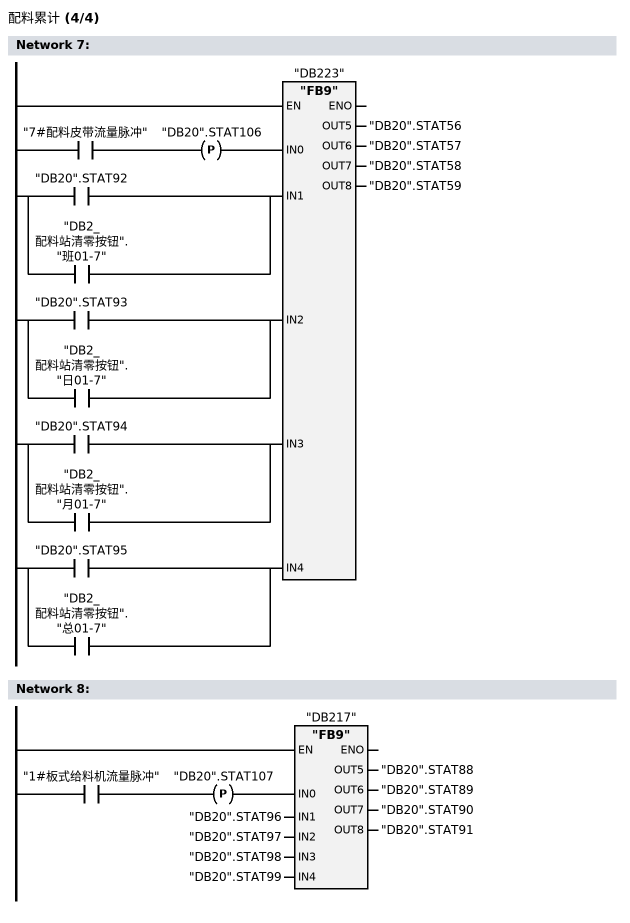
   RUNG wire#powerrail
      "DB223"(IN0 := wire#w1, IN1 := wire#w2, IN2 := wire#w3, IN3 := wire#w4, IN4 := wire#w5, OUT5 => "DB20".STAT56, OUT6 => "DB20".STAT57, OUT7 => "DB20".STAT58, OUT8 => "DB20".STAT59)
   END_RUNG
   RUNG wire#powerrail
      Contact( "7#配料皮带流量脉冲" )
      P_Trig( "DB20".STAT106 )
   END_RUNG wire#w1
   RUNG wire#powerrail
      Contact( "DB20".STAT92 )
   END_RUNG wire#w2
   RUNG wire#powerrail
      Contact( "DB2_配料站清零按钮"."班01-7" )
   END_RUNG wire#w2
   RUNG wire#powerrail
      Contact( "DB20".STAT93 )
   END_RUNG wire#w3
   RUNG wire#powerrail
      Contact( "DB2_配料站清零按钮"."日01-7" )
   END_RUNG wire#w3
   RUNG wire#powerrail
      Contact( "DB20".STAT94 )
   END_RUNG wire#w4
   RUNG wire#powerrail
      Contact( "DB2_配料站清零按钮"."月01-7" )
   END_RUNG wire#w4
   RUNG wire#powerrail
      Contact( "DB20".STAT95 )
   END_RUNG wire#w5
   RUNG wire#powerrail
      Contact( "DB2_配料站清零按钮"."总01-7" )
   END_RUNG wire#w5
   // the same network as SCL:
   #_w1 := "7#配料皮带流量脉冲" AND NOT "DB20".STAT106;   // rising edge
   "DB20".STAT106 := "7#配料皮带流量脉冲";
   "DB223"(IN0 := #_w1,   // "FB9"
           IN1 := "DB20".STAT92 OR "DB2_配料站清零按钮"."班01-7",
           IN2 := "DB20".STAT93 OR "DB2_配料站清零按钮"."日01-7",
           IN3 := "DB20".STAT94 OR "DB2_配料站清零按钮"."月01-7",
           IN4 := "DB20".STAT95 OR "DB2_配料站清零按钮"."总01-7",
           OUT5 => "DB20".STAT56,
           OUT6 => "DB20".STAT57,
           OUT7 => "DB20".STAT58,
           OUT8 => "DB20".STAT59);
END_REGION

REGION Network 8
   RUNG wire#powerrail
      "DB217"(IN0 := wire#w1, IN1 := "DB20".STAT96, IN2 := "DB20".STAT97, IN3 := "DB20".STAT98, IN4 := "DB20".STAT99, OUT5 => "DB20".STAT88, OUT6 => "DB20".STAT89, OUT7 => "DB20".STAT90, OUT8 => "DB20".STAT91)
   END_RUNG
   RUNG wire#powerrail
      Contact( "1#板式给料机流量脉冲" )
      P_Trig( "DB20".STAT107 )
   END_RUNG wire#w1
   // the same network as SCL:
   #_w1 := "1#板式给料机流量脉冲" AND NOT "DB20".STAT107;   // rising edge
   "DB20".STAT107 := "1#板式给料机流量脉冲";
   "DB217"(IN0 := #_w1,   // "FB9"
           IN1 := "DB20".STAT96,
           IN2 := "DB20".STAT97,
           IN3 := "DB20".STAT98,
           IN4 := "DB20".STAT99,
           OUT5 => "DB20".STAT88,
           OUT6 => "DB20".STAT89,
           OUT7 => "DB20".STAT90,
           OUT8 => "DB20".STAT91);
END_REGION
END_FUNCTION

FUNCTION "回转窑变频器驱动块" : Void   // FC111, LAD
{ S7_Optimized_Access := 'FALSE' }
VERSION : 0.1
   VAR_INPUT
      IN0 : Bool;   // IN0
      IN1 : Bool;   // IN1
      IN2 : Bool;   // IN2
      IN3 : Bool;   // IN3
      IN4 : Bool;   // IN4
      IN5 : Bool;   // IN5
      IN6 : Bool;   // IN6
      IN7 : Bool;   // IN7
      IN8 : Bool;   // IN8
   END_VAR
   VAR_IN_OUT
      OUT9 : Bool;   // OUT9
   END_VAR
BEGIN

REGION Network 1: OUT9
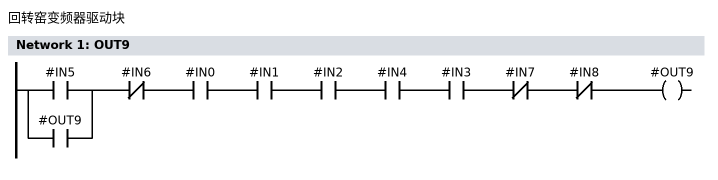
   RUNG wire#powerrail
      Contact( #IN5 )
      wire#w1
      I_Contact( #IN6 )
      Contact( #IN0 )
      Contact( #IN1 )
      Contact( #IN2 )
      Contact( #IN4 )
      Contact( #IN3 )
      I_Contact( #IN7 )
      I_Contact( #IN8 )
      Coil( #OUT9 )
   END_RUNG
   RUNG wire#powerrail
      Contact( #OUT9 )
   END_RUNG wire#w1
   // the same network as SCL:
   #OUT9 := (#IN5 OR #OUT9) AND NOT #IN6 AND #IN0 AND #IN1 AND #IN2 AND #IN4 AND #IN3 AND NOT #IN7 AND NOT #IN8;
END_REGION
END_FUNCTION

FUNCTION "回转窑接触器合闸块" : Void   // FC112, LAD
{ S7_Optimized_Access := 'FALSE' }
VERSION : 0.1
   VAR_INPUT
      IN0 : Bool;   // IN0
      IN1 : Bool;   // IN1
      IN2 : Bool;   // IN2
   END_VAR
   VAR_IN_OUT
      OUT3 : Bool;   // OUT3
   END_VAR
BEGIN

REGION Network 1: OUT3
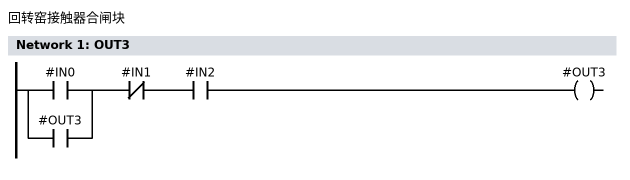
   RUNG wire#powerrail
      Contact( #IN0 )
      wire#w1
      I_Contact( #IN1 )
      Contact( #IN2 )
      Coil( #OUT3 )
   END_RUNG
   RUNG wire#powerrail
      Contact( #OUT3 )
   END_RUNG wire#w1
   // the same network as SCL:
   #OUT3 := (#IN0 OR #OUT3) AND NOT #IN1 AND #IN2;
END_REGION
END_FUNCTION

FUNCTION "稀油站功能块" : Void   // FC113, LAD
{ S7_Optimized_Access := 'FALSE' }
VERSION : 0.1
   VAR_INPUT
      LR1 : Bool;
      FAT1_1 : Bool;
      FAT1_2 : Bool;
      ST1 : Bool;
      STP1 : Bool;
      LR2 : Bool;
      FAT2_1 : Bool;
      FAT2_2 : Bool;
      ST2 : Bool;
      STP2 : Bool;
   END_VAR
   VAR_IN_OUT
      OUT10 : Bool;
      OUT11 : Bool;
   END_VAR
BEGIN

REGION Network 1
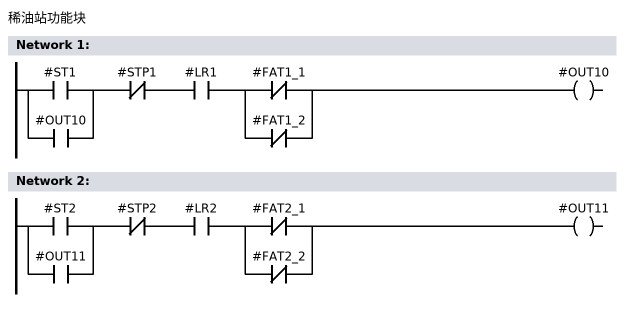
   RUNG wire#powerrail
      Contact( #ST1 )
      wire#w1
      I_Contact( #STP1 )
      Contact( #LR1 )
      wire#w2
      I_Contact( #FAT1_1 )
      wire#w3
      Coil( #OUT10 )
   END_RUNG
   RUNG wire#powerrail
      Contact( #OUT10 )
   END_RUNG wire#w1
   RUNG wire#w2
      I_Contact( #FAT1_2 )
   END_RUNG wire#w3
   // the same network as SCL:
   #OUT10 := (#ST1 OR #OUT10) AND NOT #STP1 AND #LR1 AND (NOT #FAT1_1 OR NOT #FAT1_2);
END_REGION

REGION Network 2
   RUNG wire#powerrail
      Contact( #ST2 )
      wire#w1
      I_Contact( #STP2 )
      Contact( #LR2 )
      wire#w2
      I_Contact( #FAT2_1 )
      wire#w3
      Coil( #OUT11 )
   END_RUNG
   RUNG wire#powerrail
      Contact( #OUT11 )
   END_RUNG wire#w1
   RUNG wire#w2
      I_Contact( #FAT2_2 )
   END_RUNG wire#w3
   // the same network as SCL:
   #OUT11 := (#ST2 OR #OUT11) AND NOT #STP2 AND #LR2 AND (NOT #FAT2_1 OR NOT #FAT2_2);
END_REGION
END_FUNCTION

FUNCTION "电机功能块" : Void   // FC114, LAD
{ S7_Optimized_Access := 'FALSE' }
VERSION : 0.1
   VAR_INPUT
      LR : Bool;
      FAULT : Bool;
      START : Bool;
      STOP : Bool;
   END_VAR
   VAR_IN_OUT
      OUT : Bool;
   END_VAR
BEGIN

REGION Network 1
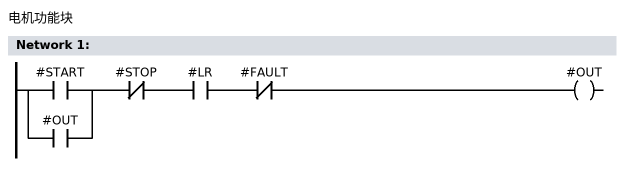
   RUNG wire#powerrail
      Contact( #START )
      wire#w1
      I_Contact( #STOP )
      Contact( #LR )
      I_Contact( #FAULT )
      Coil( #OUT )
   END_RUNG
   RUNG wire#powerrail
      Contact( #OUT )
   END_RUNG wire#w1
   // the same network as SCL:
   #OUT := (#START OR #OUT) AND NOT #STOP AND #LR AND NOT #FAULT;
END_REGION
END_FUNCTION

FUNCTION "皮带功能块" : Void   // FC115, LAD
{ S7_Optimized_Access := 'FALSE' }
VERSION : 0.1
   VAR_INPUT
      LR : Bool;
      FAULT : Bool;
      STOP : Bool;
      IN3 : Bool;
   END_VAR
   VAR_IN_OUT
      OUT : Bool;
   END_VAR
BEGIN

REGION Network 1
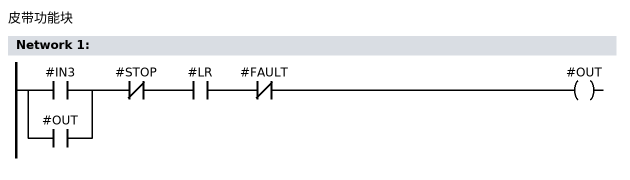
   RUNG wire#powerrail
      Contact( #IN3 )
      wire#w1
      I_Contact( #STOP )
      Contact( #LR )
      I_Contact( #FAULT )
      Coil( #OUT )
   END_RUNG
   RUNG wire#powerrail
      Contact( #OUT )
   END_RUNG wire#w1
   // the same network as SCL:
   #OUT := (#IN3 OR #OUT) AND NOT #STOP AND #LR AND NOT #FAULT;
END_REGION
END_FUNCTION

FUNCTION "脉冲累计功能块" : Void   // FC116, LAD
{ S7_Optimized_Access := 'FALSE' }
VERSION : 0.1
   VAR_INPUT
      IN0 : Bool;
      IN1 : Bool;
   END_VAR
   VAR_OUTPUT
      OUT2 : Real;
   END_VAR
   VAR_TEMP
      TEMP3 : Bool;
      TEMP4 : Real;
      TEMP5 : Real;
      TEMP6 : Real;
   END_VAR
   VAR_TEMP   // added for the SCL form of the ladder/FBD networks
      _w1 : Bool;
   END_VAR
BEGIN

REGION Network 1
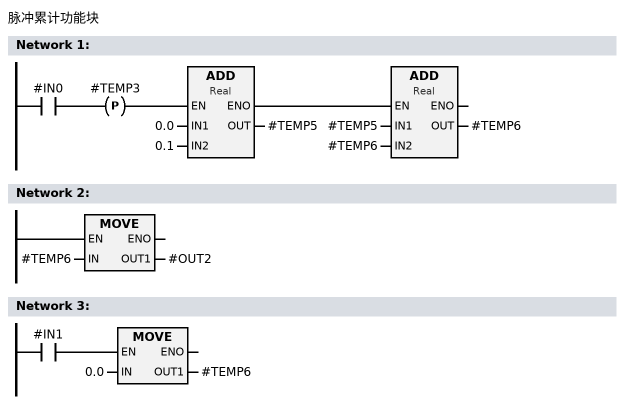
   RUNG wire#powerrail
      Contact( #IN0 )
      P_Trig( #TEMP3 )
      { S7_Templates := "SrcType := Real"; S7_GenerateENO := "TRUE" } Add(in1 := 0.0, in2 := 0.1, out => #TEMP5)
      { S7_Templates := "SrcType := Real"; S7_GenerateENO := "TRUE" } Add(in1 := #TEMP5, in2 := #TEMP6, out => #TEMP6)
   END_RUNG
   // the same network as SCL:
   // ENO of a box is taken as its EN; it also drops when the box reports an error
   #_w1 := #IN0 AND NOT #TEMP3;   // rising edge
   #TEMP3 := #IN0;
   IF #_w1 THEN
       #TEMP5 := 0.0 + 0.1;
       #TEMP6 := #TEMP5 + #TEMP6;
   END_IF;
END_REGION

REGION Network 2
   RUNG wire#powerrail
      { S7_GenerateENO := "TRUE" } Move(in := #TEMP6, out1 => #OUT2)
   END_RUNG
   // the same network as SCL:
   #OUT2 := #TEMP6;
END_REGION

REGION Network 3
   RUNG wire#powerrail
      Contact( #IN1 )
      { S7_GenerateENO := "TRUE" } Move(in := 0.0, out1 => #TEMP6)
   END_RUNG
   // the same network as SCL:
   IF #IN1 THEN #TEMP6 := 0.0; END_IF;
END_REGION

REGION Network 4 (STL)
         SET;
         SAVE;
END_REGION
END_FUNCTION

ORGANIZATION_BLOCK "Main"   // OB1, LAD, ProgramCycle
{ S7_Optimized_Access := 'FALSE' }
VERSION : 0.1
   VAR_TEMP
      TEMP0 : Byte;
      TEMP1 : Byte;
      TEMP2 : Byte;
      TEMP3 : Byte;
      TEMP4 : Byte;
      TEMP5 : Byte;
      TEMP6 : Int;
      TEMP7 : Int;
      TEMP8 : Int;
      TEMP9 : Date_And_Time;
   END_VAR
BEGIN

REGION Network 1
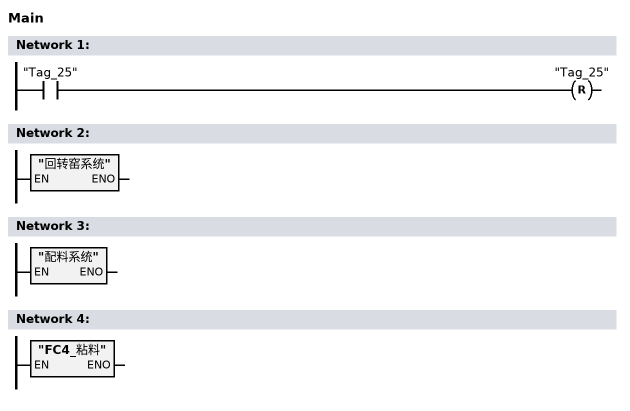
   RUNG wire#powerrail
      Contact( "Tag_25" )
      R_Coil( "Tag_25" )
   END_RUNG
   // the same network as SCL:
   IF "Tag_25" THEN "Tag_25" := FALSE; END_IF;
END_REGION

REGION Network 2
   RUNG wire#powerrail
      "回转窑系统"()
   END_RUNG
   // the same network as SCL:
   "回转窑系统"();
END_REGION

REGION Network 3
   RUNG wire#powerrail
      "配料系统"()
   END_RUNG
   // the same network as SCL:
   "配料系统"();
END_REGION

REGION Network 4
   RUNG wire#powerrail
      "FC4_粘料"()
   END_RUNG
   // the same network as SCL:
   "FC4_粘料"();
END_REGION
END_ORGANIZATION_BLOCK

ORGANIZATION_BLOCK "Cyclic interrupt"   // OB30, LAD, CyclicInterrupt
{ S7_Optimized_Access := 'TRUE' }
VERSION : 0.1
   VAR_INPUT
      Initial_Call : Bool;   // Initial call of this OB
      Event_Count : Int;   // Events discarded
   END_VAR
   VAR_TEMP   // added for the SCL form of the ladder/FBD networks
      _w1 : Bool;
      _w2 : Bool;
   END_VAR
BEGIN

REGION Network 1
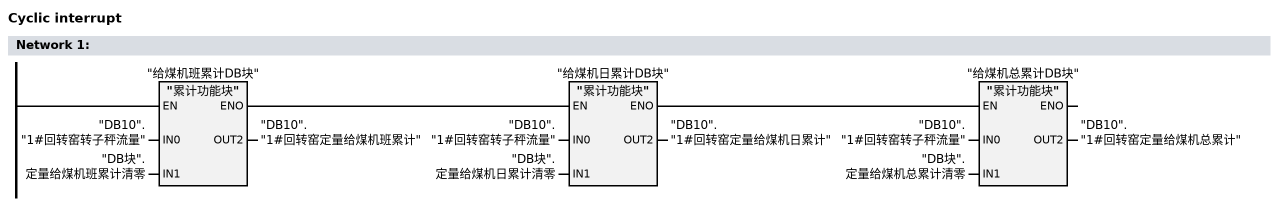
   RUNG wire#powerrail
      "给煤机班累计DB块"(IN0 := "DB10"."1#回转窑转子秤流量", IN1 := "DB块".定量给煤机班累计清零, OUT2 => "DB10"."1#回转窑定量给煤机班累计")
      "给煤机日累计DB块"(IN0 := "DB10"."1#回转窑转子秤流量", IN1 := "DB块".定量给煤机日累计清零, OUT2 => "DB10"."1#回转窑定量给煤机日累计")
      "给煤机总累计DB块"(IN0 := "DB10"."1#回转窑转子秤流量", IN1 := "DB块".定量给煤机总累计清零, OUT2 => "DB10"."1#回转窑定量给煤机总累计")
   END_RUNG
   // the same network as SCL:
   "给煤机班累计DB块"(IN0 := "DB10"."1#回转窑转子秤流量", IN1 := "DB块".定量给煤机班累计清零, OUT2 => "DB10"."1#回转窑定量给煤机班累计", ENO => #_w1);   // "累计功能块"
   "给煤机日累计DB块"(EN := #_w1,   // "累计功能块"
               IN0 := "DB10"."1#回转窑转子秤流量",
               IN1 := "DB块".定量给煤机日累计清零,
               OUT2 => "DB10"."1#回转窑定量给煤机日累计",
               ENO => #_w2);
   IF #_w2 THEN
       "给煤机总累计DB块"(IN0 := "DB10"."1#回转窑转子秤流量", IN1 := "DB块".定量给煤机总累计清零, OUT2 => "DB10"."1#回转窑定量给煤机总累计");   // "累计功能块"
   END_IF;
END_REGION
END_ORGANIZATION_BLOCK

// ===== PLC "2#DCC"  CPU 1511-1 PN =====

VAR_GLOBAL   // PLC tag table "默认变量表"
   "1#1号电场备妥" AT %I0.0 : Bool;
   "1#1号电场就绪" AT %I0.1 : Bool;
   "1#1号电场运行" AT %I0.2 : Bool;
   "1#1号电场故障" AT %I0.3 : Bool;
   "1#2号电场备妥" AT %I0.4 : Bool;
   "1#2号电场就绪" AT %I0.5 : Bool;
   "1#2号电场运行" AT %I0.6 : Bool;
   "1#2号电场故障" AT %I0.7 : Bool;
   "1#3号电场备妥" AT %I1.0 : Bool;
   "1#3号电场就绪" AT %I1.1 : Bool;
   "1#3号电场运行" AT %I1.2 : Bool;
   "1#3号电场故障" AT %I1.3 : Bool;
   "1#4号电场备妥" AT %I1.4 : Bool;
   "1#4号电场就绪" AT %I1.5 : Bool;
   "1#4号电场运行" AT %I1.6 : Bool;
   "1#4号电场故障" AT %I1.7 : Bool;
   "2#1号电场备妥" AT %I2.0 : Bool;
   "2#1号电场就绪" AT %I2.1 : Bool;
   "2#1号电场运行" AT %I2.2 : Bool;
   "2#1号电场故障" AT %I2.3 : Bool;
   "2#2号电场备妥" AT %I2.4 : Bool;
   "2#2号电场就绪" AT %I2.5 : Bool;
   "2#2号电场运行" AT %I2.6 : Bool;
   "2#2号电场故障" AT %I2.7 : Bool;
   "2#3号电场备妥" AT %I3.0 : Bool;
   "2#3号电场就绪" AT %I3.1 : Bool;
   "2#3号电场运行" AT %I3.2 : Bool;
   "2#3号电场故障" AT %I3.3 : Bool;
   "2#4号电场备妥" AT %I3.4 : Bool;
   "2#4号电场就绪" AT %I3.5 : Bool;
   "2#4号电场运行" AT %I3.6 : Bool;
   "2#4号电场故障" AT %I3.7 : Bool;
   "1#1号电场一次运行电压" AT %IW256 : Int;
   "1#1号电场一次运行电流" AT %IW258 : Int;
   "1#1号电场二次运行电压" AT %IW260 : Int;
   "1#1号电场二次运行电流" AT %IW262 : Int;
   "1#2号电场一次运行电压" AT %IW264 : Int;
   "1#2号电场一次运行电流" AT %IW266 : Int;
   "1#2号电场二次运行电压" AT %IW268 : Int;
   "1#2号电场二次运行电流" AT %IW270 : Int;
   "1#3号电场一次运行电压" AT %IW272 : Int;
   "1#3号电场一次运行电流" AT %IW274 : Int;
   "1#3号电场二次运行电压" AT %IW276 : Int;
   "1#3号电场二次运行电流" AT %IW278 : Int;
   "1#4号电场一次运行电压" AT %IW280 : Int;
   "1#4号电场一次运行电流" AT %IW282 : Int;
   "1#4号电场二次运行电压" AT %IW284 : Int;
   "1#4号电场二次运行电流" AT %IW286 : Int;
   "2#1号电场一次运行电压" AT %IW288 : Int;
   "2#1号电场一次运行电流" AT %IW290 : Int;
   "2#1号电场二次运行电压" AT %IW292 : Int;
   "2#1号电场二次运行电流" AT %IW294 : Int;
   "2#2号电场一次运行电压" AT %IW296 : Int;
   "2#2号电场一次运行电流" AT %IW298 : Int;
   "2#2号电场二次运行电压" AT %IW300 : Int;
   "2#2号电场二次运行电流" AT %IW302 : Int;
   "2#3号电场一次运行电压" AT %IW304 : Int;
   "2#3号电场一次运行电流" AT %IW306 : Int;
   "2#3号电场二次运行电压" AT %IW308 : Int;
   "2#3号电场二次运行电流" AT %IW310 : Int;
   "2#4号电场一次运行电压" AT %IW312 : Int;
   "2#4号电场一次运行电流" AT %IW314 : Int;
   "2#4号电场二次运行电压" AT %IW316 : Int;
   "2#4号电场二次运行电流" AT %IW318 : Int;
   "1#电场热风管入口压力" AT %IW320 : Int;
   "1#电场热风管出口压力" AT %IW322 : Int;
   "2#电场热风管入口压力" AT %IW324 : Int;
   "2#电场热风管出口压力" AT %IW326 : Int;
   "1#除尘热风管进口温度" AT %IW328 : Int;
   "1#除尘热风管出口温度" AT %IW330 : Int;
   "2#除尘热风管进口温度" AT %IW332 : Int;
   "2#除尘热风管出口温度" AT %IW334 : Int;
   "1#除尘U相绕组温度" AT %ID336 : Real;
   "1#除尘V相绕组温度" AT %ID340 : Real;
   "1#除尘W相绕组温度" AT %ID344 : Real;
   "1#除尘电机前轴承温度" AT %ID348 : Real;
   "1#除尘电机后轴承温度" AT %ID352 : Real;
   "1#除尘风机前轴承温度" AT %ID356 : Real;
   "1#除尘风机后轴承温度" AT %ID360 : Real;
   "2#除尘U相绕组温度" AT %ID432 : Real;
   "2#除尘V相绕组温度" AT %ID436 : Real;
   "2#除尘W相绕组温度" AT %ID440 : Real;
   "2#除尘电机前轴承温度" AT %ID444 : Real;
   "2#除尘电机后轴承温度" AT %ID448 : Real;
   "2#除尘风机前轴承温度" AT %ID452 : Real;
   "2#除尘风机后轴承温度" AT %ID456 : Real;
   "1#1号电场启动" AT %Q0.0 : Bool;
   "1#1号电场停止" AT %Q0.1 : Bool;
   "1#2号电场启动" AT %Q0.2 : Bool;
   "1#2号电场停止" AT %Q0.3 : Bool;
   "1#3号电场启动" AT %Q0.4 : Bool;
   "1#3号电场停止" AT %Q0.5 : Bool;
   "1#4号电场启动" AT %Q0.6 : Bool;
   "1#4号电场停止" AT %Q0.7 : Bool;
   "2#1号电场启动" AT %Q1.0 : Bool;
   "2#1号电场停止" AT %Q1.1 : Bool;
   "2#2号电场启动" AT %Q1.2 : Bool;
   "2#2号电场停止" AT %Q1.3 : Bool;
   "2#3号电场启动" AT %Q1.4 : Bool;
   "2#3号电场停止" AT %Q1.5 : Bool;
   "2#4号电场启动" AT %Q1.6 : Bool;
   "2#4号电场停止" AT %Q1.7 : Bool;
   "1#电除尘联锁" AT %Q2.0 : Bool;
   "2#电除尘联锁" AT %Q2.1 : Bool;
   "QB4" AT %QB4 : Byte;
   "1#1号电场控制给定" AT %QW256 : Int;
   "1#2号电场控制给定" AT %QW258 : Int;
   "1#3号电场控制给定" AT %QW260 : Int;
   "1#4号电场控制给定" AT %QW262 : Int;
   "2#1号电场控制给定" AT %QW264 : Int;
   "2#2号电场控制给定" AT %QW266 : Int;
   "2#3号电场控制给定" AT %QW268 : Int;
   "2#4号电场控制给定" AT %QW270 : Int;
   "Q2_2" AT %Q2.2 : Bool;
   "Q2_3" AT %Q2.3 : Bool;
   "Q2_4" AT %Q2.4 : Bool;
   "Q2_5" AT %Q2.5 : Bool;
   "Q2_6" AT %Q2.6 : Bool;
   "Q2_7" AT %Q2.7 : Bool;
   "Q3_0" AT %Q3.0 : Bool;
   "Q3_1" AT %Q3.1 : Bool;
   "Q3_2" AT %Q3.2 : Bool;
   "Q3_3" AT %Q3.3 : Bool;
   "Q3_4" AT %Q3.4 : Bool;
   "Q3_5" AT %Q3.5 : Bool;
   "Q3_6" AT %Q3.6 : Bool;
   "Q3_7" AT %Q3.7 : Bool;
END_VAR

DATA_BLOCK "模拟量转换DB块"   // DB1
{ S7_Optimized_Access := 'FALSE' }
VERSION : 0.1
   VAR
      "1#1号电场二次运行电压" : Real := 0.0;
      "1#1号电场二次运行电流" : Real := 0.0;
      "1#2号电场二次运行电压" : Real := 0.0;
      "1#2号电场二次运行电流" : Real := 0.0;
      "1#3号电场二次运行电压" : Real := 0.0;
      "1#3号电场二次运行电流" : Real := 0.0;
      "1#4号电场二次运行电压" : Real := 0.0;
      "1#4号电场二次运行电流" : Real := 0.0;
      "2#1号电场二次运行电压" : Real := 0.0;
      "2#1号电场二次运行电流" : Real := 0.0;
      "2#2号电场二次运行电压" : Real := 0.0;
      "2#2号电场二次运行电流" : Real := 0.0;
      "2#3号电场二次运行电压" : Real := 0.0;
      "2#3号电场二次运行电流" : Real := 0.0;
      "2#4号电场二次运行电压" : Real := 0.0;
      "2#4号电场二次运行电流" : Real := 0.0;
      "1#电场热风管入口压力" : Real := 0.0;
      "1#电场热风管出口压力" : Real := 0.0;
      "2#电场热风管入口压力" : Real := 0.0;
      "2#电场热风管出口压力" : Real := 0.0;
      "1#除尘热风管进口温度" : Real := 0.0;   // -useless
      "1#除尘热风管出口温度" : Real := 0.0;   // -useless
      "2#除尘热风管进口温度" : Real;   // -useless
      "2#除尘热风管出口温度" : Real;   // -useless
      BIPOLAR : Bool;   // 单极性，始终为0
      RET_VAL : Word := WORD#16#0000;   // 错误代码
   END_VAR
BEGIN
END_DATA_BLOCK

DATA_BLOCK "百特巡检仪温度DB块"   // DB2
{ S7_Optimized_Access := 'FALSE' }
VERSION : 0.1
   VAR
      "1#除尘U相绕组温度" : Real;   // 临时占位符变量
      "1#除尘V相绕组温度" : Real;   // 临时占位符变量
      "1#除尘W相绕组温度" : Real;   // 临时占位符变量
      "1#除尘电机前轴承温度" : Real;   // 临时占位符变量
      "1#除尘电机后轴承温度" : Real;   // 临时占位符变量
      "1#除尘风机前轴承温度" : Real;   // 临时占位符变量
      "1#除尘风机后轴承温度" : Real;   // 临时占位符变量
      DB_VAR7 : Real;   // 临时占位符变量
      DB_VAR8 : Real;   // 临时占位符变量
      DB_VAR9 : Real;   // 临时占位符变量
      DB_VAR10 : Real;   // 临时占位符变量
      DB_VAR11 : Real;   // 临时占位符变量
      DB_VAR12 : Real;   // 临时占位符变量
      DB_VAR13 : Real;   // 临时占位符变量
      DB_VAR14 : Real;   // 临时占位符变量
      DB_VAR15 : Real;   // 临时占位符变量
      DB_VAR16 : Real;   // 临时占位符变量
      DB_VAR17 : Real;   // 临时占位符变量
      DB_VAR18 : Real;   // 临时占位符变量
      DB_VAR19 : Real;   // 临时占位符变量
      DB_VAR20 : Real;   // 临时占位符变量
      DB_VAR21 : Real;   // 临时占位符变量
      DB_VAR22 : Real;   // 临时占位符变量
      DB_VAR23 : Real;   // 临时占位符变量
      DB_VAR24 : Real;   // 临时占位符变量
      DB_VAR25 : Real;   // 临时占位符变量
      DB_VAR26 : Real;   // 临时占位符变量
      DB_VAR27 : Real;   // 临时占位符变量
      DB_VAR28 : Real;   // 临时占位符变量
      DB_VAR29 : Real;   // 临时占位符变量
      DB_VAR30 : Real;   // 临时占位符变量
      DB_VAR31 : Real;   // 临时占位符变量
      DB_VAR32 : Real;   // 临时占位符变量
      DB_VAR33 : Real;   // 临时占位符变量
      DB_VAR34 : Real;   // 临时占位符变量
      DB_VAR35 : Real;   // 临时占位符变量
      DB_VAR36 : Real;   // 临时占位符变量
      DB_VAR37 : Real;   // 临时占位符变量
      DB_VAR38 : Real;   // 临时占位符变量
      DB_VAR39 : Real;   // 临时占位符变量
      DB_VAR40 : Real;   // 临时占位符变量
      DB_VAR41 : Real;   // 临时占位符变量
      DB_VAR42 : Real;   // 临时占位符变量
      DB_VAR43 : Real;   // 临时占位符变量
      DB_VAR44 : Real;   // 临时占位符变量
      DB_VAR45 : Real;   // 临时占位符变量
      DB_VAR46 : Real;   // 临时占位符变量
      DB_VAR47 : Real;   // 临时占位符变量
      DB_VAR48 : Real;   // 临时占位符变量
      DB_VAR49 : Real;   // 临时占位符变量
      "2#除尘U相绕组温度" : Real;   // 临时占位符变量
      "2#除尘V相绕组温度" : Real;   // 临时占位符变量
      "2#除尘W相绕组温度" : Real;   // 临时占位符变量
      "2#除尘电机前轴承温度" : Real;   // 临时占位符变量
      "2#除尘电机后轴承温度" : Real;   // 临时占位符变量
      "2#除尘风机前轴承温度" : Real;   // 临时占位符变量
      "2#除尘风机后轴承温度" : Real;   // 临时占位符变量
      DB_VAR57 : Real;   // 临时占位符变量
      DB_VAR58 : Real;   // 临时占位符变量
      DB_VAR59 : Real;   // 临时占位符变量
      DB_VAR60 : Real;   // 临时占位符变量
      DB_VAR61 : Real;   // 临时占位符变量
      DB_VAR62 : Real;   // 临时占位符变量
      DB_VAR63 : Real;   // 临时占位符变量
      DB_VAR64 : Real;   // 临时占位符变量
      DB_VAR65 : Real;   // 临时占位符变量
      DB_VAR66 : Real;   // 临时占位符变量
   END_VAR
BEGIN
END_DATA_BLOCK

FUNCTION "FC1" : Void   // FC1, LAD
{ S7_Optimized_Access := 'FALSE' }
VERSION : 0.1
BEGIN

REGION Network 1: 1#1号电场二次运行电压
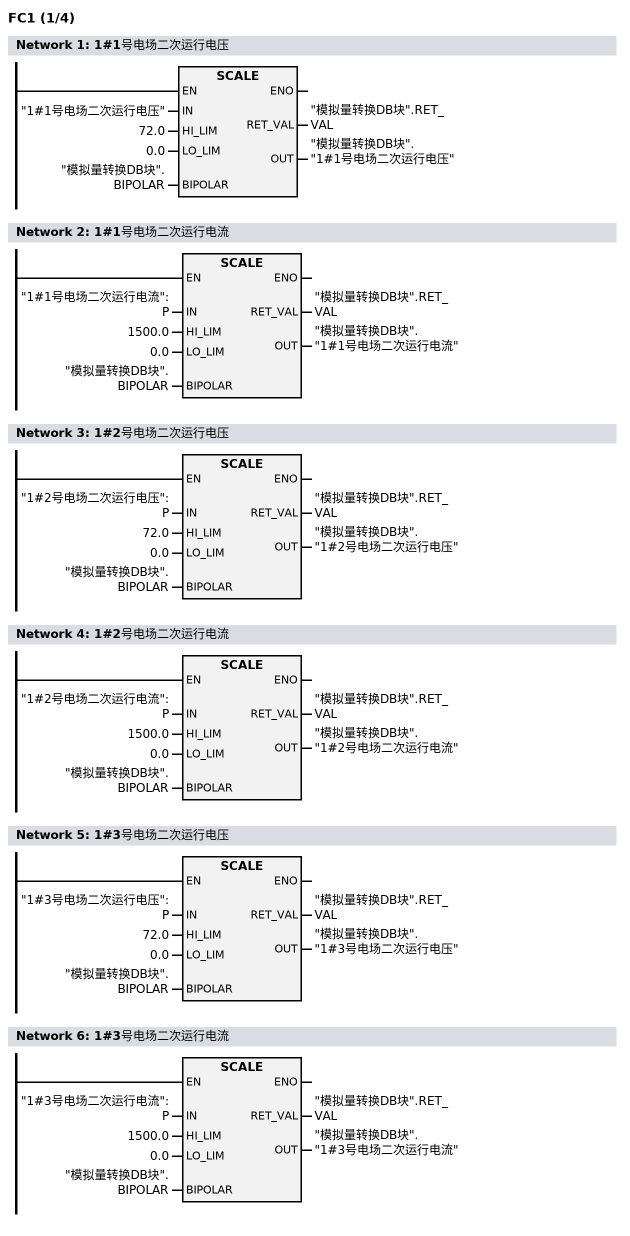
   "模拟量转换DB块".RET_VAL := SCALE(IN := "1#1号电场二次运行电压",
                           HI_LIM := 72.0,
                           LO_LIM := 0.0,
                           BIPOLAR := "模拟量转换DB块".BIPOLAR,
                           OUT => "模拟量转换DB块"."1#1号电场二次运行电压");
END_REGION

REGION Network 2: 1#1号电场二次运行电流
   "模拟量转换DB块".RET_VAL := SCALE(IN := "1#1号电场二次运行电流":P,
                           HI_LIM := 1500.0,
                           LO_LIM := 0.0,
                           BIPOLAR := "模拟量转换DB块".BIPOLAR,
                           OUT => "模拟量转换DB块"."1#1号电场二次运行电流");
END_REGION

REGION Network 3: 1#2号电场二次运行电压
   "模拟量转换DB块".RET_VAL := SCALE(IN := "1#2号电场二次运行电压":P,
                           HI_LIM := 72.0,
                           LO_LIM := 0.0,
                           BIPOLAR := "模拟量转换DB块".BIPOLAR,
                           OUT => "模拟量转换DB块"."1#2号电场二次运行电压");
END_REGION

REGION Network 4: 1#2号电场二次运行电流
   "模拟量转换DB块".RET_VAL := SCALE(IN := "1#2号电场二次运行电流":P,
                           HI_LIM := 1500.0,
                           LO_LIM := 0.0,
                           BIPOLAR := "模拟量转换DB块".BIPOLAR,
                           OUT => "模拟量转换DB块"."1#2号电场二次运行电流");
END_REGION

REGION Network 5: 1#3号电场二次运行电压
   "模拟量转换DB块".RET_VAL := SCALE(IN := "1#3号电场二次运行电压":P,
                           HI_LIM := 72.0,
                           LO_LIM := 0.0,
                           BIPOLAR := "模拟量转换DB块".BIPOLAR,
                           OUT => "模拟量转换DB块"."1#3号电场二次运行电压");
END_REGION

REGION Network 6: 1#3号电场二次运行电流
   "模拟量转换DB块".RET_VAL := SCALE(IN := "1#3号电场二次运行电流":P,
                           HI_LIM := 1500.0,
                           LO_LIM := 0.0,
                           BIPOLAR := "模拟量转换DB块".BIPOLAR,
                           OUT => "模拟量转换DB块"."1#3号电场二次运行电流");
END_REGION

REGION Network 7: 1#4号电场二次运行电压
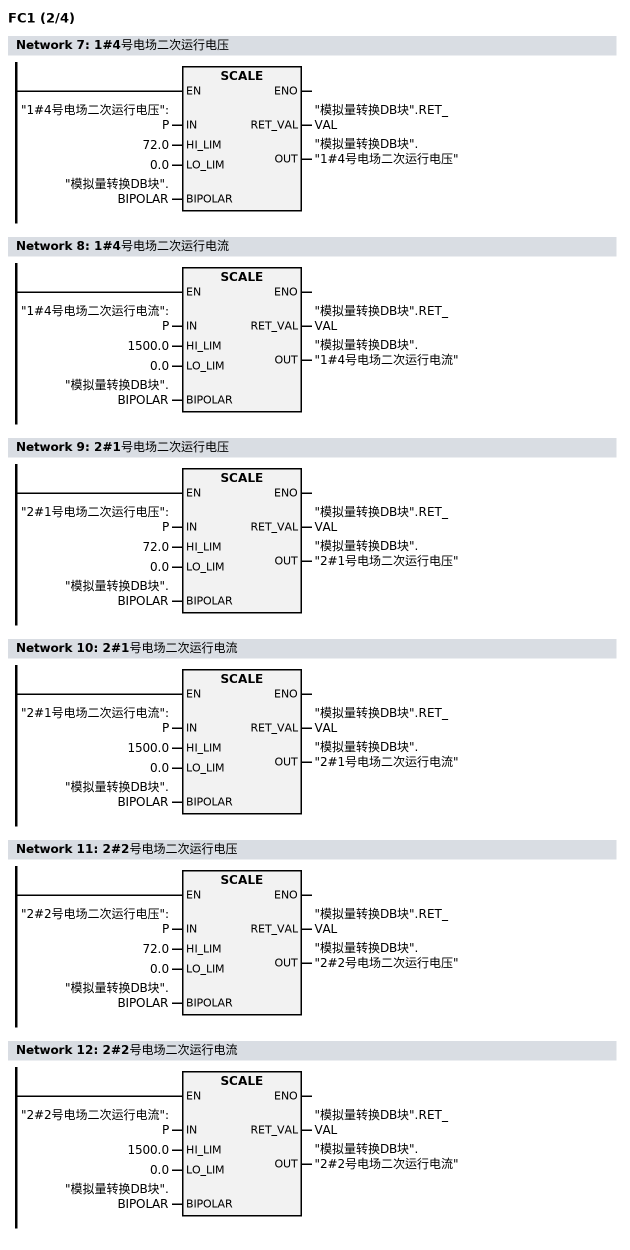
   "模拟量转换DB块".RET_VAL := SCALE(IN := "1#4号电场二次运行电压":P,
                           HI_LIM := 72.0,
                           LO_LIM := 0.0,
                           BIPOLAR := "模拟量转换DB块".BIPOLAR,
                           OUT => "模拟量转换DB块"."1#4号电场二次运行电压");
END_REGION

REGION Network 8: 1#4号电场二次运行电流
   "模拟量转换DB块".RET_VAL := SCALE(IN := "1#4号电场二次运行电流":P,
                           HI_LIM := 1500.0,
                           LO_LIM := 0.0,
                           BIPOLAR := "模拟量转换DB块".BIPOLAR,
                           OUT => "模拟量转换DB块"."1#4号电场二次运行电流");
END_REGION

REGION Network 9: 2#1号电场二次运行电压
   "模拟量转换DB块".RET_VAL := SCALE(IN := "2#1号电场二次运行电压":P,
                           HI_LIM := 72.0,
                           LO_LIM := 0.0,
                           BIPOLAR := "模拟量转换DB块".BIPOLAR,
                           OUT => "模拟量转换DB块"."2#1号电场二次运行电压");
END_REGION

REGION Network 10: 2#1号电场二次运行电流
   "模拟量转换DB块".RET_VAL := SCALE(IN := "2#1号电场二次运行电流":P,
                           HI_LIM := 1500.0,
                           LO_LIM := 0.0,
                           BIPOLAR := "模拟量转换DB块".BIPOLAR,
                           OUT => "模拟量转换DB块"."2#1号电场二次运行电流");
END_REGION

REGION Network 11: 2#2号电场二次运行电压
   "模拟量转换DB块".RET_VAL := SCALE(IN := "2#2号电场二次运行电压":P,
                           HI_LIM := 72.0,
                           LO_LIM := 0.0,
                           BIPOLAR := "模拟量转换DB块".BIPOLAR,
                           OUT => "模拟量转换DB块"."2#2号电场二次运行电压");
END_REGION

REGION Network 12: 2#2号电场二次运行电流
   "模拟量转换DB块".RET_VAL := SCALE(IN := "2#2号电场二次运行电流":P,
                           HI_LIM := 1500.0,
                           LO_LIM := 0.0,
                           BIPOLAR := "模拟量转换DB块".BIPOLAR,
                           OUT => "模拟量转换DB块"."2#2号电场二次运行电流");
END_REGION

REGION Network 13: 2#3号电场二次运行电压
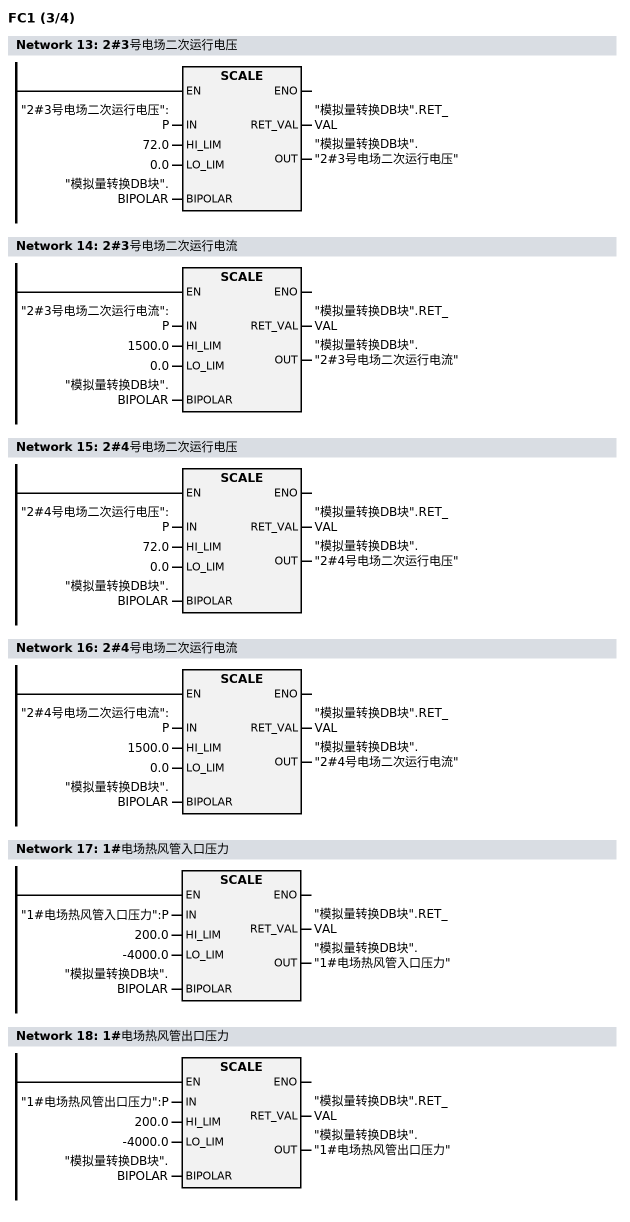
   "模拟量转换DB块".RET_VAL := SCALE(IN := "2#3号电场二次运行电压":P,
                           HI_LIM := 72.0,
                           LO_LIM := 0.0,
                           BIPOLAR := "模拟量转换DB块".BIPOLAR,
                           OUT => "模拟量转换DB块"."2#3号电场二次运行电压");
END_REGION

REGION Network 14: 2#3号电场二次运行电流
   "模拟量转换DB块".RET_VAL := SCALE(IN := "2#3号电场二次运行电流":P,
                           HI_LIM := 1500.0,
                           LO_LIM := 0.0,
                           BIPOLAR := "模拟量转换DB块".BIPOLAR,
                           OUT => "模拟量转换DB块"."2#3号电场二次运行电流");
END_REGION

REGION Network 15: 2#4号电场二次运行电压
   "模拟量转换DB块".RET_VAL := SCALE(IN := "2#4号电场二次运行电压":P,
                           HI_LIM := 72.0,
                           LO_LIM := 0.0,
                           BIPOLAR := "模拟量转换DB块".BIPOLAR,
                           OUT => "模拟量转换DB块"."2#4号电场二次运行电压");
END_REGION

REGION Network 16: 2#4号电场二次运行电流
   "模拟量转换DB块".RET_VAL := SCALE(IN := "2#4号电场二次运行电流":P,
                           HI_LIM := 1500.0,
                           LO_LIM := 0.0,
                           BIPOLAR := "模拟量转换DB块".BIPOLAR,
                           OUT => "模拟量转换DB块"."2#4号电场二次运行电流");
END_REGION

REGION Network 17: 1#电场热风管入口压力
   "模拟量转换DB块".RET_VAL := SCALE(IN := "1#电场热风管入口压力":P,
                           HI_LIM := 200.0,
                           LO_LIM := -4000.0,
                           BIPOLAR := "模拟量转换DB块".BIPOLAR,
                           OUT => "模拟量转换DB块"."1#电场热风管入口压力");
END_REGION

REGION Network 18: 1#电场热风管出口压力
   "模拟量转换DB块".RET_VAL := SCALE(IN := "1#电场热风管出口压力":P,
                           HI_LIM := 200.0,
                           LO_LIM := -4000.0,
                           BIPOLAR := "模拟量转换DB块".BIPOLAR,
                           OUT => "模拟量转换DB块"."1#电场热风管出口压力");
END_REGION

REGION Network 19: 2#电场热风管入口压力
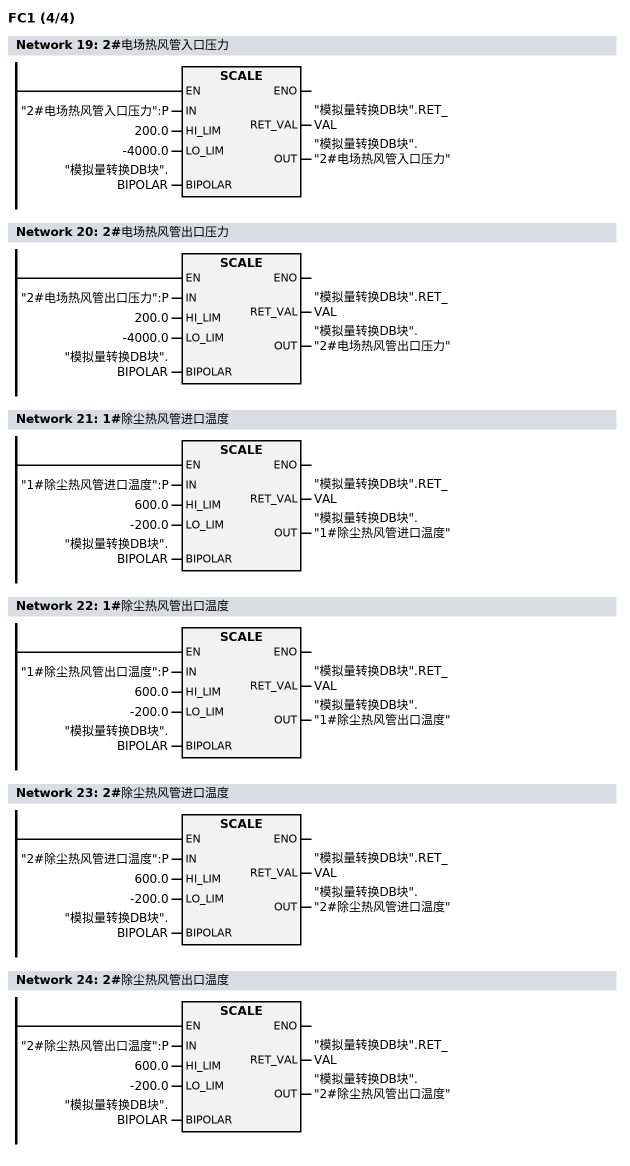
   "模拟量转换DB块".RET_VAL := SCALE(IN := "2#电场热风管入口压力":P,
                           HI_LIM := 200.0,
                           LO_LIM := -4000.0,
                           BIPOLAR := "模拟量转换DB块".BIPOLAR,
                           OUT => "模拟量转换DB块"."2#电场热风管入口压力");
END_REGION

REGION Network 20: 2#电场热风管出口压力
   "模拟量转换DB块".RET_VAL := SCALE(IN := "2#电场热风管出口压力":P,
                           HI_LIM := 200.0,
                           LO_LIM := -4000.0,
                           BIPOLAR := "模拟量转换DB块".BIPOLAR,
                           OUT => "模拟量转换DB块"."2#电场热风管出口压力");
END_REGION

REGION Network 21: 1#除尘热风管进口温度
   "模拟量转换DB块".RET_VAL := SCALE(IN := "1#除尘热风管进口温度":P,
                           HI_LIM := 600.0,
                           LO_LIM := -200.0,
                           BIPOLAR := "模拟量转换DB块".BIPOLAR,
                           OUT => "模拟量转换DB块"."1#除尘热风管进口温度");
END_REGION

REGION Network 22: 1#除尘热风管出口温度
   "模拟量转换DB块".RET_VAL := SCALE(IN := "1#除尘热风管出口温度":P,
                           HI_LIM := 600.0,
                           LO_LIM := -200.0,
                           BIPOLAR := "模拟量转换DB块".BIPOLAR,
                           OUT => "模拟量转换DB块"."1#除尘热风管出口温度");
END_REGION

REGION Network 23: 2#除尘热风管进口温度
   "模拟量转换DB块".RET_VAL := SCALE(IN := "2#除尘热风管进口温度":P,
                           HI_LIM := 600.0,
                           LO_LIM := -200.0,
                           BIPOLAR := "模拟量转换DB块".BIPOLAR,
                           OUT => "模拟量转换DB块"."2#除尘热风管进口温度");
END_REGION

REGION Network 24: 2#除尘热风管出口温度
   "模拟量转换DB块".RET_VAL := SCALE(IN := "2#除尘热风管出口温度":P,
                           HI_LIM := 600.0,
                           LO_LIM := -200.0,
                           BIPOLAR := "模拟量转换DB块".BIPOLAR,
                           OUT => "模拟量转换DB块"."2#除尘热风管出口温度");
END_REGION
END_FUNCTION

FUNCTION "DP&MODBUS通讯" : Void   // FC15, LAD
{ S7_Optimized_Access := 'FALSE' }
VERSION : 0.1
BEGIN

REGION Network 1
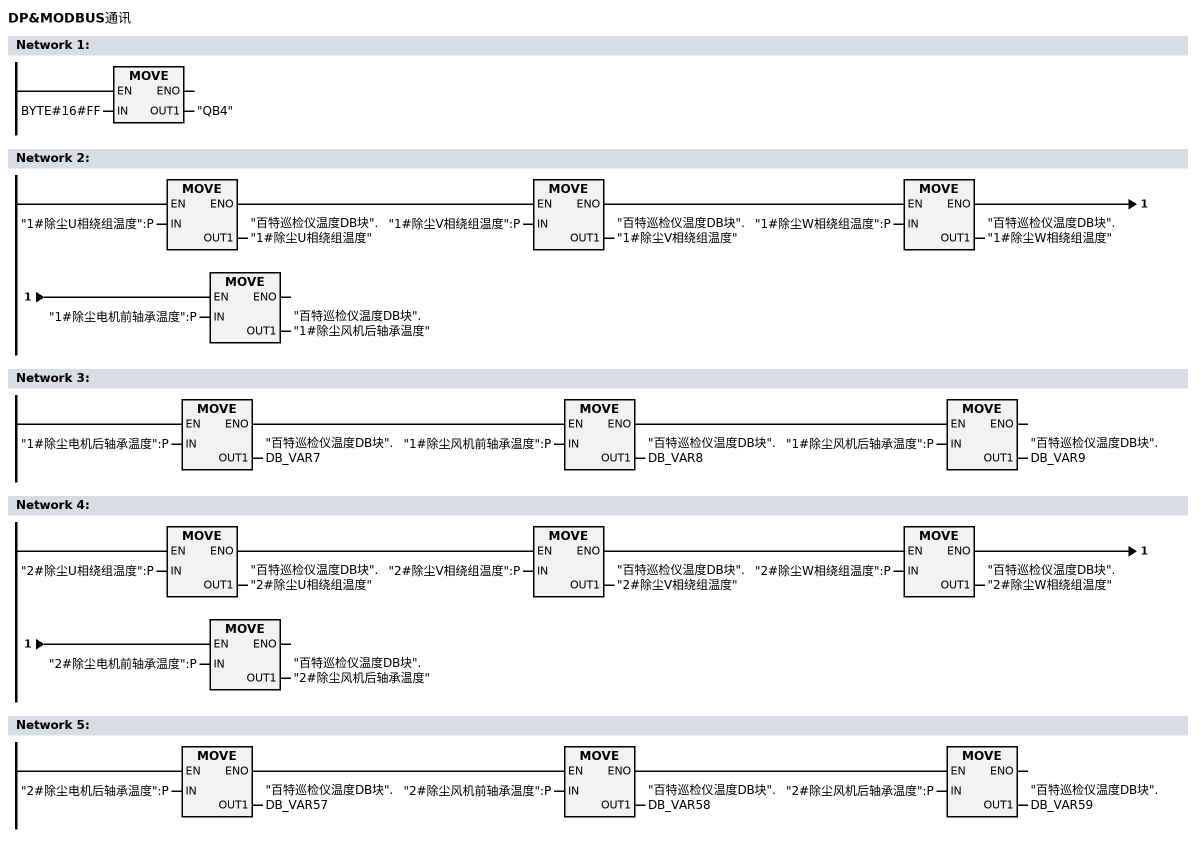
   RUNG wire#powerrail
      { S7_GenerateENO := "TRUE" } Move(in := BYTE#16#FF, out1 => "QB4")
   END_RUNG
   // the same network as SCL:
   "QB4" := BYTE#16#FF;
END_REGION

REGION Network 2
   RUNG wire#powerrail
      { S7_GenerateENO := "TRUE" } Move(in := "1#除尘U相绕组温度":P, out1 => "百特巡检仪温度DB块"."1#除尘U相绕组温度")
      { S7_GenerateENO := "TRUE" } Move(in := "1#除尘V相绕组温度":P, out1 => "百特巡检仪温度DB块"."1#除尘V相绕组温度")
      { S7_GenerateENO := "TRUE" } Move(in := "1#除尘W相绕组温度":P, out1 => "百特巡检仪温度DB块"."1#除尘W相绕组温度")
      { S7_GenerateENO := "TRUE" } Move(in := "1#除尘电机前轴承温度":P, out1 => "百特巡检仪温度DB块"."1#除尘风机后轴承温度")
   END_RUNG
   // the same network as SCL:
   // ENO of a box is taken as its EN; it also drops when the box reports an error
   "百特巡检仪温度DB块"."1#除尘U相绕组温度" := "1#除尘U相绕组温度":P;
   "百特巡检仪温度DB块"."1#除尘V相绕组温度" := "1#除尘V相绕组温度":P;
   "百特巡检仪温度DB块"."1#除尘W相绕组温度" := "1#除尘W相绕组温度":P;
   "百特巡检仪温度DB块"."1#除尘风机后轴承温度" := "1#除尘电机前轴承温度":P;
END_REGION

REGION Network 3
   RUNG wire#powerrail
      { S7_GenerateENO := "TRUE" } Move(in := "1#除尘电机后轴承温度":P, out1 => "百特巡检仪温度DB块".DB_VAR7)
      { S7_GenerateENO := "TRUE" } Move(in := "1#除尘风机前轴承温度":P, out1 => "百特巡检仪温度DB块".DB_VAR8)
      { S7_GenerateENO := "TRUE" } Move(in := "1#除尘风机后轴承温度":P, out1 => "百特巡检仪温度DB块".DB_VAR9)
   END_RUNG
   // the same network as SCL:
   // ENO of a box is taken as its EN; it also drops when the box reports an error
   "百特巡检仪温度DB块".DB_VAR7 := "1#除尘电机后轴承温度":P;
   "百特巡检仪温度DB块".DB_VAR8 := "1#除尘风机前轴承温度":P;
   "百特巡检仪温度DB块".DB_VAR9 := "1#除尘风机后轴承温度":P;
END_REGION

REGION Network 4
   RUNG wire#powerrail
      { S7_GenerateENO := "TRUE" } Move(in := "2#除尘U相绕组温度":P, out1 => "百特巡检仪温度DB块"."2#除尘U相绕组温度")
      { S7_GenerateENO := "TRUE" } Move(in := "2#除尘V相绕组温度":P, out1 => "百特巡检仪温度DB块"."2#除尘V相绕组温度")
      { S7_GenerateENO := "TRUE" } Move(in := "2#除尘W相绕组温度":P, out1 => "百特巡检仪温度DB块"."2#除尘W相绕组温度")
      { S7_GenerateENO := "TRUE" } Move(in := "2#除尘电机前轴承温度":P, out1 => "百特巡检仪温度DB块"."2#除尘风机后轴承温度")
   END_RUNG
   // the same network as SCL:
   // ENO of a box is taken as its EN; it also drops when the box reports an error
   "百特巡检仪温度DB块"."2#除尘U相绕组温度" := "2#除尘U相绕组温度":P;
   "百特巡检仪温度DB块"."2#除尘V相绕组温度" := "2#除尘V相绕组温度":P;
   "百特巡检仪温度DB块"."2#除尘W相绕组温度" := "2#除尘W相绕组温度":P;
   "百特巡检仪温度DB块"."2#除尘风机后轴承温度" := "2#除尘电机前轴承温度":P;
END_REGION

REGION Network 5
   RUNG wire#powerrail
      { S7_GenerateENO := "TRUE" } Move(in := "2#除尘电机后轴承温度":P, out1 => "百特巡检仪温度DB块".DB_VAR57)
      { S7_GenerateENO := "TRUE" } Move(in := "2#除尘风机前轴承温度":P, out1 => "百特巡检仪温度DB块".DB_VAR58)
      { S7_GenerateENO := "TRUE" } Move(in := "2#除尘风机后轴承温度":P, out1 => "百特巡检仪温度DB块".DB_VAR59)
   END_RUNG
   // the same network as SCL:
   // ENO of a box is taken as its EN; it also drops when the box reports an error
   "百特巡检仪温度DB块".DB_VAR57 := "2#除尘电机后轴承温度":P;
   "百特巡检仪温度DB块".DB_VAR58 := "2#除尘风机前轴承温度":P;
   "百特巡检仪温度DB块".DB_VAR59 := "2#除尘风机后轴承温度":P;
END_REGION
END_FUNCTION

ORGANIZATION_BLOCK "Main"   // OB1, LAD, ProgramCycle
TITLE = "Main Program Sweep (Cycle)"
{ S7_Optimized_Access := 'TRUE' }
VERSION : 0.1
   VAR_INPUT
      Initial_Call : Bool;   // Initial call of this OB
      Remanence : Bool;   // =True, if remanent data are available
   END_VAR
BEGIN

REGION Network 1
